// Mitsubishi GX Works2 project: 40国轩高温2次注液尝试优化   PLC: Q06UDEH

TYPE ConveyorIO : STRUCT
  xUnloadCCW : BOOL;  (* 下料为反转 *)
  xUnloadAlarm : BOOL;  (* 下料报警 *)
  xUnload : BOOL;  (* 下料请求 *)
  xPutInto : BOOL;  (* 线体直接投入物料 *)
  xNotArriveAlarm : BOOL;  (* 未到达报警 *)
  xNextRun : BOOL;  (* 下段线体运行 *)
  xMotorCW : BOOL;  (* 电机正转 *)
  xMotorCCW : BOOL;  (* 电机反转 *)
  xManual : BOOL;  (* 手动 *)
  xloadCCW : BOOL;  (* 上料为反转 *)
  xLimitAlarrm : BOOL;  (* 限位报警 *)
  xLoad : BOOL;  (* 上料请求 *)
  xForward : BOOL;  (* 正转手动 *)
  xEmpty : BOOL;  (* 线体状态为空 *)
  xCWPresent : BOOL;  (* 正转检测有无传感器 *)
  xCCWPresent : BOOL;  (* 反转检测有无传感器 *)
  xBusy : BOOL;  (* 工作中 *)
  xBackward : BOOL;  (* 反转手动 *)
  xAuto : BOOL;  (* 自动 *)
  xPosLimit : BOOL;  (* 正限位 *)
  xNegLimit : BOOL;  (* 负限位 *)
  xOverWidthAlarm : BOOL;  (* 超宽报警 *)
  xError : BOOL;  (* 报警 *)
  iProductCategoryIn : INT;  (* 产品类型输入 *)
  iProductCategory : INT;  (* 产品类型记录 *)
  iProductCategoryOut : INT;  (* 产品类型输出 *)
  diDeviceID : DINT;  (* 设备编号 *)
  tUnloadAlarmDelay : TIME;  (* 下料报警时间设置 *)
  tLoadDelay : TIME;  (* 上料延时设置 *)
  xSizeDeficientDetect : BOOL;  (* 尺寸缺陷检测 *)
  xZoneClear : BOOL;  (* 初始化线体清除 *)
  tZoneClearTime : TIME;  (* 初始化线体清除时间 *)
  iTaskIDIn : INT;  (* 产品类型输入 *)
  iTaskID : INT;  (* 产品类型记录 *)
  iTaskIDOut : INT;  (* 产品类型输出 *)
  diDesConveyorIn : DINT;  (* 产品类型输入 *)
  diDesConveyor : DINT;  (* 产品类型记录 *)
  diDesConveyorOut : DINT;  (* 产品类型输出 *)
END_STRUCT END_TYPE

TYPE ShuttleCarIO : STRUCT
  xReady : BOOL;  (* 准备就绪 *)
  xForward : BOOL;  (* 正转 *)
  xBackward : BOOL;  (* 反转 *)
  iCurrentPos : INT;  (* 当前位置 *)
  iDestinationPos : INT;  (* 目标位置 *)
  xCW : BOOL;  (* 正转输出 *)
  xCCW : BOOL;  (* 反转输出 *)
  xBrake : BOOL;  (* 刹车 *)
  xHomeSwitch : BOOL;  (* 零位接近开关 *)
  xPosLimit : BOOL;  (* 正限位 *)
  xNegLimit : BOOL;  (* 负限位 *)
  xMDIExe : BOOL;  (* MDI开始 *)
  xMDIDone : BOOL;  (* MDI 完成 *)
  xPassLimit : BOOL;  (* 限位屏蔽 *)
  xPosLimitCatch : BOOL;  (* 正限位捕捉 *)
  xNegLimitCatch : BOOL;  (* 负限位捕捉 *)
  xHomeExe : BOOL;  (* 开始寻零 *)
  xHomeDone : BOOL;  (* 寻零完成 *)
  xHomeBusy : BOOL;  (* 寻零中 *)
  xHomeFailed : BOOL;  (* 寻零失败 *)
  xBusy : BOOL;  (* 工作中 *)
  tArriveDelay : TIME;  (* 到位延时 *)
  xCylinder : BOOL;  (* 气缸控制 *)
  tBrakeDelay : TIME;  (* 抱闸延时 *)
  xPauseRamp : BOOL;  (* 暂停减速斜坡标志位 *)
  xPresentDetect1 : BOOL;  (* 物料有无检测1 *)
  xPresentDetect2 : BOOL;  (* 物料有无检测2 *)
  xOvertimeAlarm : BOOL;  (* 超时报警 *)
  tSetOverTime : TIME;  (* 设置超时时间 *)
  xLooseDetect : BOOL;  (* 松绳检测 *)
  xLooseAlarm : BOOL;  (* 松绳报警 *)
  xArrive : BOOL;  (* 到位信号 *)
  diDeviceID : DINT;  (* 设备编号 *)
  xMoveStep : BOOL;  (* 寸动 *)
  xAdrSwitch : ARRAY [1..8] OF BOOL;  (* 位置开关 *)
END_STRUCT END_TYPE

TYPE SwitchIO : STRUCT
  xLiftCylinderRetractDetect : BOOL;
  xLiftCylinderExtendDetect : BOOL;
  xLiftCylinderRetract : BOOL;
  xLiftCylinderExtend : BOOL;
  xEntryBarCylinderRetract : BOOL;
  xLiftCylinderExtendInit : BOOL;
  xEntryEnable : BOOL;
  xExitEnable : BOOL;
  xExitBarCylinderRetract : BOOL;
  xSwithEnable : BOOL;
  xLiftCylinderRetractButton : BOOL;
  xLiftCylinderExtendButton : BOOL;
  xEntryBarCylinderRetractButton : BOOL;
  xExitBarCylinderRetractButton : BOOL;
  xPutInto : BOOL;  (* 单体复位 *)
  tSetOvertime : TIME;  (* 设定超时报警时间 *)
  xOvertimeAlarm : BOOL;  (* 超时报警 *)
END_STRUCT END_TYPE

TYPE QueueElement : STRUCT
  xCondition : BOOL;
  iPriority : INT;
END_STRUCT END_TYPE

TYPE UConveyorIO : STRUCT
  xLiftCylinderRetractDetect1 : BOOL;
  xLiftCylinderRetractDetect2 : BOOL;
  xLiftCylinderExtendDetect1 : BOOL;
  xLiftCylinderExtendDetect2 : BOOL;
  xLiftCylinderRetract1 : BOOL;
  xLiftCylinderRetract2 : BOOL;
  xLiftCylinderExtend1 : BOOL;
  xLiftCylinderExtend2 : BOOL;
  xExitBarCylinderRetract1 : BOOL;
  xExitBarCylinderRetract2 : BOOL;
  xLiftCylinderExtendInit1 : BOOL;
  xLiftCylinderExtendInit2 : BOOL;
  xEntryEnable1 : BOOL;
  xEntryEnable2 : BOOL;
  xEntryEnable3 : BOOL;
  xExitEnable1 : BOOL;
  xExitEnable2 : BOOL;
  xExitEnable3 : BOOL;
  xPassEnable : BOOL;  (* 直接放行去下段 *)
  xLiftCylinderRetractButton1 : BOOL;
  xLiftCylinderRetractButton2 : BOOL;
  xLiftCylinderExtendButton1 : BOOL;
  xLiftCylinderExtendButton2 : BOOL;
  xExitBarCylinderRetractButton1 : BOOL;
  xExitBarCylinderRetractButton2 : BOOL;
  xPutInto : BOOL;  (* 单体复位 *)
  tSetOvertime : TIME;  (* 设定超时报警时间 *)
  xOvertimeAlarm : BOOL;  (* 超时报警 *)
  iTask : INT;  (* 3个任务 *)
  xBatteryDetect1 : BOOL;  (* 电池检测1 *)
  xBatteryDetect2 : BOOL;  (* 电池检测2 *)
  xBatteryError : BOOL;  (* 空框里有电池错误 *)
END_STRUCT END_TYPE

TYPE FolderIO : STRUCT
  o_xCylinderGrabExtend : BOOL;  (* 气缸夹紧 *)
  o_xCylinderGrabRetract : BOOL;  (* 气缸松开 *)
  i_xCylinderGrabExtendDetect : BOOL;  (* 夹紧检测 *)
  i_xCylinderGrabRetractDetect : BOOL;  (* 松开检测 *)
  o_xCylinderUpExtend : BOOL;  (* 上层伸出 *)
  o_xCylinderUpRetract : BOOL;  (* 上层缩回 *)
  i_xCylinderUpExtendDetect : BOOL;  (* 上层伸出检测 *)
  i_xCylinderUpRetractDetect : BOOL;  (* 上层缩回检测 *)
  o_xCylinderDownExtend : BOOL;  (* 下层伸出 *)
  o_xCylinderDownRetract : BOOL;  (* 下层缩回 *)
  i_xCylinderDownExtendDetect : BOOL;  (* 下层伸出检测 *)
  i_xCylinderDownRetractDetect : BOOL;  (* 下层缩回检测 *)
  i_xExitEnable : BOOL;  (* 下料信号 *)
  i_xEntryEnable : BOOL;  (* 上料信号 *)
  o_xEntryPermit : BOOL;  (* 允许上料(拆盘需要，叠盘不需要) *)
  i_iFloor : INT;  (* 层数 *)
  i_xCylinderGrabExtendButton : BOOL;  (* 气缸夹紧按钮 *)
  i_xCylinderGrabRetractButton : BOOL;  (* 气缸松开按钮 *)
  i_xCylinderUpExtendButton : BOOL;  (* 上层伸出按钮 *)
  i_xCylinderUpRetractButton : BOOL;  (* 上层缩回按钮 *)
  i_xCylinderDownExtendButton : BOOL;  (* 下层伸出按钮 *)
  i_xCylinderDownRetractButton : BOOL;  (* 下层缩回按钮 *)
  o_xDownCylinderError : BOOL;  (* 下层气缸层伸出未到达 *)
  o_xUpCylinderError : BOOL;  (* 上层气缸伸出未到达 *)
  o_xGrabCylinderError : BOOL;  (* 夹紧气缸伸出未到达 *)
  i_tSetOvertime : TIME;  (* 未到达计时 *)
END_STRUCT END_TYPE

TYPE CommunicationIO : STRUCT
  i_iResponsPCPLC : INT;  (* 上位机写入-请求确认 *)
  i_iTypeInfoPCPLC : INT;  (* 上位机写入-批次标识，是否同批次 *)
  i_iReadWriteFlagPCPLC : INT;  (* 上位机写入-读写标志位 *)
  i_iTaskProcessFlagPCPLC : INT;  (* 上位机写入-任务处理标志位 *)
  i_iCommandPCPLC : INT;  (* 上位机写入-命令字 *)
  i_iTaskIDPCPLC : INT;  (* 上位机写入-任务号 *)
  i_diDestinationDevicePCPLC : DINT;  (* 上位机写入-目标设备号 *)
  i_iProductIDPCPLC : INT;  (* 上位机写入-框码后4位 *)
  o_iRequestPLCPC : INT;  (* 上位机读取-请求状态 *)
  o_iForceInportPLCPC : INT;  (* 上位机读取-强制入库 *)
  o_iFolderNumberPLCPC : INT;  (* 上位机读取-叠盘数量 *)
  o_iEmptyPLCPC : INT;  (* 上位机读取-有料状态 *)
  o_iReadWriteFlagPLCPC : INT;  (* 上位机读取-读写标志位 *)
  o_iDeviceStatusPLCPC : INT;  (* 上位机读取-设备状态 *)
  o_iTaskIDPLCPC : INT;  (* 上位机读取-任务号 *)
  o_iProductIDPLCPC : INT;  (* 上位机读取-框码后4位 *)
  i_xExtraCondition : BOOL;  (* 发送请求时的额外条件,比如需要升降到位 *)
  i_xExportConveyor : BOOL;  (* 线体是出库线体还是入库线体 *)
  i_xImportConveyor : BOOL;  (* 入库线体 *)
END_STRUCT END_TYPE

// global labels: Global
VAR_GLOBAL
  g_xAuto AT M11 : BOOL;
  g_xAutoSwitch AT X1 : BOOL;  (* 手自动钥匙旋钮 *)
  g_xManual : BOOL;
  g_xEStop AT X0 : BOOL;
  g_xAlarm : BOOL;
  g_xMute : BOOL;
  g_xStackLampRed AT Y200 : BOOL;
  g_xStackLampAmber AT Y201 : BOOL;
  g_xStackLampGreen AT Y202 : BOOL;
  g_xStop AT X3 : BOOL;
  g_xPause AT M3 : BOOL;  (* 暂停 *)
  g_xAutoStart AT X2 : BOOL;
  g_xAutoLamp AT Y204 : BOOL;
  g_xRemoteAutoStart AT M0 : BOOL;
  g_iConveyorStatus AT D4 : INT;
  g_xBuzzer AT Y203 : BOOL;
  g_xRemoteAuto AT M10 : BOOL;
  g_xReset AT X4 : BOOL;
  g_xResetSingle AT M4 : BOOL;  (* 单线体复位 *)
  g_xInsertTask AT M5 : BOOL;  (* 插入任务 *)
  g_diInsertDesConveyor AT D8 : DINT;
  g_iInsertTaskID AT D2 : INT;  (* 插入任务号 *)
  g_iInsertCategory AT D6 : INT;
  g_iState AT D40 : INT;
  g_iLocalAutoStep : BOOL;
  g_diDeviceIDSelect AT D0 : DINT;
  g_xTcpFailed : BOOL;  (* 通讯失败 *)
  g_xPickOver : ARRAY [1..4] OF BOOL;  (* 注液机给我们的信号，待定 *)
  g_x36HourExport1Forbidden AT M2 : BOOL;  (* 36H出库禁止 *)
  g_xForceImport AT M1 : BOOL;  (* 强制入库 *)
END_VAR

// task Task_01 (event TRUE, interval 0, priority 31): POU, START, TCP

PROGRAM POU
VAR
  Conveyor40102 : Conveyor;
  Conveyor40104 : Conveyor;
  Conveyor40105 : Conveyor;
  Conveyor40106 : Conveyor;
  Conveyor40103 : Conveyor;
  Conveyor40107 : Conveyor;
  Conveyor40108 : Conveyor;
  Conveyor40101 : Conveyor;
  Conveyor40109 : Conveyor;
  Conveyor40110 : Conveyor;
  Conveyor40111 : Conveyor;
  Conveyor40113 : Conveyor;
  Conveyor40114 : Conveyor;
  Conveyor40115 : Conveyor;
  Conveyor40116 : Conveyor;
  Conveyor40117 : Conveyor;
  Conveyor40118 : Conveyor;
  Conveyor40119 : Conveyor;
  Conveyor40120 : Conveyor;
  Conveyor40122 : Conveyor;
  Conveyor40124 : Conveyor;
  Conveyor40126 : Conveyor;
  Conveyor40129 : Conveyor;
  Conveyor40131 : Conveyor;
  Conveyor40133 : Conveyor;
  Conveyor40136 : Conveyor;
  Conveyor40137 : Conveyor;
  Conveyor40138 : Conveyor;
  Conveyor40140 : Conveyor;
  Conveyor401021 : Conveyor;
  Conveyor401101 : Conveyor;
  ConveyorIO40101 : ConveyorIO;
  ConveyorIO40103 : ConveyorIO;
  ConveyorIO40104 : ConveyorIO;
  ConveyorIO40105 : ConveyorIO;
  ConveyorIO40106 : ConveyorIO;
  ConveyorIO40107 : ConveyorIO;
  ConveyorIO40108 : ConveyorIO;
  ConveyorIO40109 : ConveyorIO;
  ConveyorIO40110 : ConveyorIO;
  ConveyorIO40111 : ConveyorIO;
  ConveyorIO40112 : ConveyorIO;
  ConveyorIO40113 : ConveyorIO;
  ConveyorIO40114 : ConveyorIO;
  ConveyorIO40115 : ConveyorIO;
  ConveyorIO40116 : ConveyorIO;
  ConveyorIO40117 : ConveyorIO;
  ConveyorIO40118 : ConveyorIO;
  ConveyorIO40119 : ConveyorIO;
  ConveyorIO40122 : ConveyorIO;
  ConveyorIO40124 : ConveyorIO;
  ConveyorIO40126 : ConveyorIO;
  ConveyorIO40128 : ConveyorIO;
  ConveyorIO40131 : ConveyorIO;
  ConveyorIO40132 : ConveyorIO;
  ConveyorIO40133 : ConveyorIO;
  ConveyorIO40135 : ConveyorIO;
  ConveyorIO40136 : ConveyorIO;
  ConveyorIO40137 : ConveyorIO;
  ConveyorIO40140 : ConveyorIO;
  ConveyorIO401021 : ConveyorIO;
  ConveyorIO401101 : ConveyorIO;
  Lifter40202 : ShuttleCar;
  Lifter40203 : ShuttleCar;
  Lifter40204 : ShuttleCar;
  Lifter40206 : ShuttleCar;
  LifterIO40202 : ShuttleCarIO;
  LifterIO40203 : ShuttleCarIO;
  LifterIO40204 : ShuttleCarIO;
  LifterIO40206 : ShuttleCarIO;
  Switch40302 : Switch;
  Switch40303 : Switch;
  Switch40304 : Switch;
  Switch40306 : Switch;
  Switch40307 : Switch;
  Switch40308 : Switch;
  Switch40309 : Switch;
  SwitchIO40301 : SwitchIO;
  SwitchIO40302 : SwitchIO;
  SwitchIO40303 : SwitchIO;
  SwitchIO40304 : SwitchIO;
  SwitchIO40305 : SwitchIO;
  SwitchIO40306 : SwitchIO;
  SwitchIO40307 : SwitchIO;
  SwitchIO40308 : SwitchIO;
  SwitchIO40309 : SwitchIO;
  Folder40501 : Folder;
  FolderIO40501 : FolderIO;
  DivideFolder40502 : DivideFolder;
  DivideFolderIO40502 : FolderIO;
  ConveyorIO40129 : ConveyorIO;
  Conveyor40112 : Conveyor;
  ConveyorIO40138 : ConveyorIO;
  Conveyor40128 : Conveyor;
  Conveyor40135 : Conveyor;
  Conveyor401061 : Conveyor;
  Lifter40201 : ShuttleCar;
  LifterIO40201 : ShuttleCarIO;
  Switch40301 : Switch;
  Conveyor40132 : Conveyor;
  ConveyorIO40102 : ConveyorIO;
  ConveyorIO401061 : ConveyorIO;
  Lifter40205 : ShuttleCar;
  LifterIO40205 : ShuttleCarIO;
  Switch40305 : Switch;
  Switch40310 : Switch;
  Switch40311 : Switch;
  Switch40312 : Switch;
  SwitchIO40310 : SwitchIO;
  SwitchIO40311 : SwitchIO;
  SwitchIO40312 : SwitchIO;
  ComConveyor40140 : ConveyorCommunication;
  ComConveyor40209 : ConveyorCommunication;
  ComConveyor40111 : ConveyorCommunication;
  ComConveyor40104 : ConveyorCommunication;
  ComConveyor40105 : ConveyorCommunication;
  ComConveyorIO40140 : CommunicationIO;
  ComConveyorIO40209 : CommunicationIO;
  ComConveyorIO40111 : CommunicationIO;
  ComConveyorIO40104 : CommunicationIO;
  ComConveyorIO40105 : CommunicationIO;
  Task40105 : PriorityQueue;  (* 4个位置要料请求排队 *)
  TaskCondition40105 : ARRAY [1..13] OF QueueElement;  (* 4个位置要料请求排队 *)
  m_iTask40105 : INT;  (* 4个位置要料请求排队 *)
  m_xLoadPermit : ARRAY [1..4] OF BOOL;  (* 4个·位置的上料许可，用触摸屏控制 *)
  m_xPickStrat : ARRAY [1..4] OF BOOL;  (* 4个位置的开始取料信号，给到注液机器 *)
  m_xPickDone : ARRAY [1..4] OF BOOL;  (* 4个取料完毕信号，注液机给我们 *)
  Conveyor401131 : Conveyor;
  Conveyor401161 : Conveyor;
  Conveyor401191 : Conveyor;
  ConveyorIO40120 : ConveyorIO;
  ConveyorIO401161 : ConveyorIO;
  ConveyorIO401131 : ConveyorIO;
  ConveyorIO401191 : ConveyorIO;
  Lifter40207 : ShuttleCar;
  Lifter40208 : ShuttleCar;
  LifterIO40207 : ShuttleCarIO;
  LifterIO40208 : ShuttleCarIO;
  Conveyor40134 : Conveyor;
  ConveyorIO40134 : ConveyorIO;
  ConveyorIO40209 : ConveyorIO;
  Conveyor40209 : Conveyor;
  m_xImport : BOOL;  (* 高温房上料多转一会儿 *)
  m_xExport : BOOL;  (* 高温房下料多转一会儿 *)
  m_TonImportDelay : TON;  (* 高温房入库延时 *)
  m_xImportDelay : BOOL;  (* 高温房入库延时 *)
  m_tImportDelay : TIME;  (* 高温房入库延时 *)
  m_TonExportDelay : TON;  (* 高温房出库延时 *)
  m_xExportDelay : BOOL;  (* 高温房出库延时 *)
  m_tExportDelay : TIME;  (* 高温房出库延时 *)
  TaskSwitch40305 : PreemptivePriority;  (* 1线入口任务队列 *)
  TaskCondition40305 : ARRAY [1..13] OF BOOL;  (* 1线入口任务队列 *)
  m_iTask40305 : INT;  (* 1线入口任务队列 *)
  TaskSwitch40306 : PreemptivePriority;  (* 2线入口任务队列 *)
  TaskCondition40306 : ARRAY [1..13] OF BOOL;  (* 2线入口任务队列 *)
  m_iTask40306 : INT;  (* 2线入口任务队列 *)
  TaskSwitch40307 : PreemptivePriority;  (* 3线入口任务队列 *)
  TaskCondition40307 : ARRAY [1..13] OF BOOL;  (* 3线入口任务队列 *)
  m_iTask40307 : INT;  (* 3线入口任务队列 *)
END_VAR
(*与注液机对接信号*)(*
	Y205:=M700;
	Y206:=M701;
	Y207:=M702;
	Y239:=M703;
	M705:=X4A AND X4B AND X4C AND X4D;
	*)
	OUT_T(m_xPickStrat[1] AND g_xAuto , TC1 ,10 );
	OUT_T(m_xPickStrat[2] AND g_xAuto , TC2 ,10 );
	OUT_T(m_xPickStrat[3] AND g_xAuto , TC3 ,10 );
	OUT_T(m_xPickStrat[4] AND g_xAuto , TC4 ,10 );
	Y205:=TS1;(*他们要求到位延时1秒给信号*)
	Y206:=TS2;
	Y207:=TS3;
	Y239:=TS4;
	g_xPickOver[1]:=X4A;
	g_xPickOver[2]:=X4B;
	g_xPickOver[3]:=X4C;
	g_xPickOver[4]:=X4D;		
Conveyor40140(ConveyorMotor:=ConveyorIO40140);(*叠盘前，虚拟扫码工位*)														
ConveyorIO40140.diDeviceID:=40140;	
ConveyorIO40140.xCWPresent:=D421.7;(*不良品工位的光电*)
ConveyorIO40140.xPutInto:=D421.9;(*状态刷新*)

Conveyor40209(ConveyorMotor:=ConveyorIO40209);(*起始叠盘和高温入横向线体*)
ConveyorIO40209.xCWPresent:=X39;						
Y234:=ConveyorIO40209.xMotorCW OR ConveyorIO40101.xMotorCW;						
ConveyorIO40209.xForward:=M542;						
M339:= NOT ConveyorIO40209.xEmpty;						
M639:=ConveyorIO40209.xError;						
ConveyorIO40209.diDeviceID:=40209;	
ConveyorIO40209.tLoadDelay:=t#4000ms;

Conveyor40101(ConveyorMotor:=ConveyorIO40101);(*高温入库横向*)
ConveyorIO40101.xCWPresent:=X8;						
(*Y208:=ConveyorIO40101.xMotorCW;						
ConveyorIO40101.xForward:=M500;*)						
M301:= NOT ConveyorIO40101.xEmpty;						
M601:=ConveyorIO40101.xError;						
ConveyorIO40101.diDeviceID:=40101;						
ConveyorIO40101.tLoadDelay:=t#4000ms;

Conveyor40102(ConveyorMotor:=ConveyorIO40102);(*高温入库竖向*)
ConveyorIO40102.xCCWPresent:=X8;
Y209:=ConveyorIO40102.xMotorCW OR ConveyorIO401021.xMotorCW;						
ConveyorIO40102.xForward:=M501;						
M302:= NOT ConveyorIO401021.xEmpty;						
M602:=ConveyorIO40102.xError OR ConveyorIO401021.xError;						
ConveyorIO40102.diDeviceID:=401021;						

Conveyor401021(ConveyorMotor:=ConveyorIO401021);(*虚拟的，入库门前停止位*)
ConveyorIO401021.xCWPresent:=X9;						
ConveyorIO401021.diDeviceID:=40102;		

Conveyor40103(ConveyorMotor:=ConveyorIO40103);(*高温入库门后，竖向*)
ConveyorIO40103.xCWPresent:=XA OR X5;					
Y20A:=ConveyorIO40103.xMotorCW;						
ConveyorIO40103.xForward:=M502;						
M303:= NOT ConveyorIO40103.xEmpty;						
M603:=ConveyorIO40103.xError;						
ConveyorIO40103.diDeviceID:=40103;						
ConveyorIO40103.tLoadDelay:=t#4000ms;

Conveyor40104(ConveyorMotor:=ConveyorIO40104);(*高温入库后横向*)
ConveyorIO40104.xCWPresent:=XA OR X5;						
Y20B:=ConveyorIO40104.xMotorCW OR m_xImport;						
ConveyorIO40104.xForward:=M503;						
M304:= NOT ConveyorIO40104.xEmpty;						
M604:=ConveyorIO40104.xError;						
ConveyorIO40104.diDeviceID:=40104;	

Conveyor40111(ConveyorMotor:=ConveyorIO40111);(*高温入库对接线体*)										
ConveyorIO40111.xCWPresent:=X7E;						
Y212:=ConveyorIO40111.xMotorCW;						
ConveyorIO40111.xForward:=M510;						
M311:= NOT ConveyorIO40111.xEmpty;						
M611:=ConveyorIO40111.xError;						
ConveyorIO40111.diDeviceID:=40111;	
ConveyorIO40111.tLoadDelay:=t#2S;	

Conveyor40105(ConveyorMotor:=ConveyorIO40105);(*高温出库对接线体*)
ConveyorIO40105.xCWPresent:=X7B;						
Y20C:=ConveyorIO40105.xMotorCW;						
ConveyorIO40105.xForward:=M504;						
M305:= NOT ConveyorIO40105.xEmpty;						
M605:=ConveyorIO40105.xError;						
ConveyorIO40105.diDeviceID:=40105;						

Conveyor40108(ConveyorMotor:=ConveyorIO40108);(*高温出库里面横向*)
ConveyorIO40108.xCWPresent:=XF OR X7;						
Y20F:=ConveyorIO40108.xMotorCW OR m_xExport;						
ConveyorIO40108.xForward:=M507;						
M308:= NOT ConveyorIO40108.xEmpty;						
M608:=ConveyorIO40108.xError;						
ConveyorIO40108.diDeviceID:=40108;	
ConveyorIO40108.tLoadDelay:=T#4000MS;

Conveyor40107(ConveyorMotor:=ConveyorIO40107);(*高温出库，里面竖向*)
ConveyorIO40107.xCWPresent:=XF OR X7;						
Y20E:=ConveyorIO40107.xMotorCW OR ConveyorIO401061.xMotorCW;						
ConveyorIO40107.xForward:=M506;						
M307:= NOT ConveyorIO401061.xEmpty;						
M607:=ConveyorIO40107.xError OR ConveyorIO401061.xError;						
ConveyorIO40107.diDeviceID:=401061;		

Conveyor401061(ConveyorMotor:=ConveyorIO401061);(*出库门前停止位，虚拟一段*)
ConveyorIO401061.xCWPresent:=XE;										
ConveyorIO401061.diDeviceID:=40107;	

Conveyor40106(ConveyorMotor:=ConveyorIO40106);(*高温出库，外面竖向*)
ConveyorIO40106.xCWPresent:=XD;						
Y20D:=ConveyorIO40106.xMotorCW;						
ConveyorIO40106.xForward:=M505;						
M306:= NOT ConveyorIO40106.xEmpty;						
M606:=ConveyorIO40106.xError;						
ConveyorIO40106.diDeviceID:=40106;															
ConveyorIO40106.tLoadDelay:=T#4000MS;

Conveyor40109(ConveyorMotor:=ConveyorIO40109);(*高温出库横向,&拆盘机&1线横向*)
ConveyorIO40109.xCWPresent:=XD;						
Y224:=ConveyorIO40109.xMotorCW OR ConveyorIO40117.xMotorCW OR ConveyorIO40114.xMotorCW;						
ConveyorIO40109.xForward:=M508;						
M309:= NOT ConveyorIO40109.xEmpty;						
M609:=ConveyorIO40109.xError;						
ConveyorIO40109.diDeviceID:=40109;		

Conveyor40117(ConveyorMotor:=ConveyorIO40117);(*拆盘位置*)					
ConveyorIO40117.xCWPresent:=XC;									
ConveyorIO40117.xForward:=M516;						
M317:= NOT ConveyorIO40117.xEmpty;						
M617:=ConveyorIO40117.xError;						
ConveyorIO40117.diDeviceID:=40117;
ConveyorIO40117.tLoadDelay:=t#4000ms;

Conveyor40114(ConveyorMotor:=ConveyorIO40114);(*1线横向*)					
ConveyorIO40114.xCWPresent:=X10;											
M314:= NOT ConveyorIO40114.xEmpty;						
M614:=ConveyorIO40114.xError;						
ConveyorIO40114.diDeviceID:=40114;						
ConveyorIO40114.tLoadDelay:=T#2000MS;

Conveyor40110(ConveyorMotor:=ConveyorIO40110);(*1线入*)
ConveyorIO40110.xCWPresent:=X10;						
Y211:=ConveyorIO40110.xMotorCW OR ConveyorIO401101.xMotorCW;						
ConveyorIO40110.xForward:=M509;								
M610:=ConveyorIO40110.xError OR ConveyorIO401101.xError;						
ConveyorIO40110.diDeviceID:=401101;					

Conveyor401101(ConveyorMotor:=ConveyorIO401101);(*1线末端*)
ConveyorIO401101.xPosLimit:= X88;
ConveyorIO401101.xNegLimit:=X89;
ConveyorIO401101.xCWPresent:=X12;											
M310:= NOT ConveyorIO401101.xEmpty;			
ConveyorIO401101.diDeviceID:=40110;	
ConveyorIO401101.tLoadDelay:=t#1000ms;
Y278:=(g_xAuto AND NOT ConveyorIO401101.xEmpty AND NOT m_xPickDone[1] AND NOT M585)(*夹紧气缸*)
			OR(g_xManual AND M585);		(*AND NOT M585 临时这么改一下，因为他们测试阶段，需要人工拿走托盘，就要松开夹紧气缸*)
Y27F:=ConveyorIO401101.xNextRun OR (g_xManual AND M586);(*末端阻挡*)		

Conveyor40112(ConveyorMotor:=ConveyorIO40112);(*2线横向*)
ConveyorIO40112.xCWPresent:=X13;						
Y213:=ConveyorIO40112.xMotorCW;						
ConveyorIO40112.xForward:=M511;						
M312:= NOT ConveyorIO40112.xEmpty;						
M612:=ConveyorIO40112.xError;						
ConveyorIO40112.diDeviceID:=40112;						
ConveyorIO40112.tLoadDelay:=T#7500MS;


Conveyor40113(ConveyorMotor:=ConveyorIO40113);(*2线入*)
ConveyorIO40113.xCWPresent:=X13;						
Y214:=ConveyorIO40113.xMotorCW OR ConveyorIO401131.xMotorCW;						
ConveyorIO40113.xForward:=M512;											
M613:=ConveyorIO40113.xError OR ConveyorIO401131.xError;						
ConveyorIO40113.diDeviceID:=401131;										

Conveyor401131(ConveyorMotor:=ConveyorIO401131);(*2线末端*)
ConveyorIO401131.xPosLimit:= X8A;
ConveyorIO401131.xNegLimit:=X8B;
ConveyorIO401131.xCWPresent:=X15;											
M313:= NOT ConveyorIO401131.xEmpty;											
ConveyorIO401131.diDeviceID:=40113;	
ConveyorIO401131.tLoadDelay:=t#1000ms;
Y272:=(g_xAuto AND NOT ConveyorIO401131.xEmpty AND NOT m_xPickDone[2] AND NOT M587)(*夹紧气缸*)
			OR(g_xManual AND M587);		(*AND NOT M587 临时这么改一下，因为他们测试阶段，需要人工拿走托盘，就要松开夹紧气缸*)	
Y27E:=ConveyorIO401131.xNextRun OR (g_xManual AND M588);(*末端阻挡*)			

Conveyor40115(ConveyorMotor:=ConveyorIO40115);(*3线横向*)
ConveyorIO40115.xCWPresent:=X16;						
Y216:=ConveyorIO40115.xMotorCW;						
ConveyorIO40115.xForward:=M514;						
M315:= NOT ConveyorIO40115.xEmpty;						
M615:=ConveyorIO40115.xError;						
ConveyorIO40115.diDeviceID:=40115;						
ConveyorIO40115.tLoadDelay:=T#5000MS;

Conveyor40116(ConveyorMotor:=ConveyorIO40116)(*3线入*);
ConveyorIO40116.xCWPresent:=X16;						
Y217:=ConveyorIO40116.xMotorCW OR ConveyorIO401161.xMotorCW;						
ConveyorIO40116.xForward:=M515;											
M616:=ConveyorIO40116.xError OR ConveyorIO401161.xError;						
ConveyorIO40116.diDeviceID:=401161;								

Conveyor401161(ConveyorMotor:=ConveyorIO401161)(*3线末端*);
ConveyorIO401161.xPosLimit:=X8C;
ConveyorIO401191.xNegLimit:=X8D;
ConveyorIO401161.xCWPresent:=X18;									
M316:= NOT ConveyorIO401161.xEmpty;										
ConveyorIO401161.diDeviceID:=40116;	
ConveyorIO401161.tLoadDelay:=t#1000ms;
Y27D:=(g_xAuto AND NOT ConveyorIO401161.xEmpty AND NOT m_xPickDone[3] AND NOT M589)(*夹紧气缸*)
			OR(g_xManual AND M589);		(*AND NOT M587 临时这么改一下，因为他们测试阶段，需要人工拿走托盘，就要松开夹紧气缸*)	
Y274:=ConveyorIO401161.xNextRun OR (g_xManual AND M590);(*末端阻挡*)	

Conveyor40118(ConveyorMotor:=ConveyorIO40118);(*4线横向**)
ConveyorIO40118.xCWPresent:=X19;						
Y219:=ConveyorIO40118.xMotorCW;						
ConveyorIO40118.xForward:=M517;						
M318:= NOT ConveyorIO40118.xEmpty;						
M618:=ConveyorIO40118.xError;						
ConveyorIO40118.diDeviceID:=40118;						
ConveyorIO40118.tLoadDelay:=T#4000MS;

Conveyor40119(ConveyorMotor:=ConveyorIO40119);(*4线入*)
ConveyorIO40119.xCWPresent:=X19;						
Y21A:=ConveyorIO40119.xMotorCW OR ConveyorIO401191.xMotorCW;						
ConveyorIO40119.xForward:=M518;											
M619:=ConveyorIO40119.xError OR ConveyorIO40119.xError;						
ConveyorIO40119.diDeviceID:=401191;						

Conveyor401191(ConveyorMotor:=ConveyorIO401191);(*4线末端*)
ConveyorIO401191.xPosLimit:=1(*X1B*);
ConveyorIO401191.xNegLimit:=X93;
ConveyorIO401191.xCWPresent:=X92;											
M319:= NOT ConveyorIO401191.xEmpty;											
ConveyorIO401191.diDeviceID:=40119;
ConveyorIO401191.tLoadDelay:=t#1000ms;	
Y27C:=(g_xAuto AND NOT ConveyorIO401191.xEmpty AND NOT m_xPickDone[4] AND NOT M591)(*夹紧气缸*)
			OR(g_xManual AND M591);		(*AND NOT M587 临时这么改一下，因为他们测试阶段，需要人工拿走托盘，就要松开夹紧气缸*)	
Y245:=ConveyorIO401191.xNextRun OR (g_xManual AND M592);(*末端阻挡*)	


Conveyor40120(ConveyorMotor:=ConveyorIO40120);(*下层4横*)
(*ConveyorIO40120.xPosLimit:=X92;						
ConveyorIO40120.xNegLimit:=X93;		*)				
ConveyorIO40120.xCWPresent:=X1D;						
Y21E:=ConveyorIO40120.xMotorCW;						
ConveyorIO40120.xForward:=M519;						
M320:= NOT ConveyorIO40120.xEmpty;						
M620:=ConveyorIO40120.xError;						
ConveyorIO40120.diDeviceID:=40120;						
(*
Conveyor40121(ConveyorMotor:=ConveyorIO40121);
ConveyorIO40121.xCWPresent:=X1C;						
Y21C:=ConveyorIO40121.xMotorCW;						
ConveyorIO40121.xForward:=M520;						
M321:= NOT ConveyorIO40121.xEmpty;						
M621:=ConveyorIO40121.xError;						
ConveyorIO40121.diDeviceID:=40121;						
*)
Conveyor40122(ConveyorMotor:=ConveyorIO40122);(*下层4出*)
ConveyorIO40122.xCWPresent:=X1D;						
Y21D:=ConveyorIO40122.xMotorCW;						
ConveyorIO40122.xForward:=M521;						
M322:= NOT ConveyorIO40122.xEmpty;						
M622:=ConveyorIO40122.xError;						
ConveyorIO40122.diDeviceID:=40122;		
ConveyorIO40122.tLoadDelay:=T#4000MS;				
(*
Conveyor40123(ConveyorMotor:=ConveyorIO40123);
ConveyorIO40123.xCWPresent:=X1D;						
Y21E:=ConveyorIO40123.xMotorCW;						
ConveyorIO40123.xForward:=M522;						
M323:= NOT ConveyorIO40123.xEmpty;						
M623:=ConveyorIO40123.xError;						
ConveyorIO40123.diDeviceID:=40123;		*)				

Conveyor40124(ConveyorMotor:=ConveyorIO40124);(*下层3出*)
ConveyorIO40124.xCWPresent:=X20;						
Y21F:=ConveyorIO40124.xMotorCW;						
ConveyorIO40124.xForward:=M523;						
M324:= NOT ConveyorIO40124.xEmpty;						
M624:=ConveyorIO40124.xError;						
ConveyorIO40124.diDeviceID:=40124;		
ConveyorIO40124.tLoadDelay:=T#4000MS;				
(*
Conveyor40125(ConveyorMotor:=ConveyorIO40125);
ConveyorIO40125.xCWPresent:=X20;						
Y220:=ConveyorIO40125.xMotorCW;						
ConveyorIO40125.xForward:=M524;						
M325:= NOT ConveyorIO40125.xEmpty;						
M625:=ConveyorIO40125.xError;						
ConveyorIO40125.diDeviceID:=40125;						
*)
Conveyor40126(ConveyorMotor:=ConveyorIO40126);(*下层3横*)
ConveyorIO40126.xCWPresent:=X20;						
Y221:=ConveyorIO40126.xMotorCW;						
ConveyorIO40126.xForward:=M525;						
M326:= NOT ConveyorIO40126.xEmpty;						
M626:=ConveyorIO40126.xError;						
ConveyorIO40126.diDeviceID:=40126;									

Conveyor40128(ConveyorMotor:=ConveyorIO40128);(*下层2出*)
ConveyorIO40128.xCWPresent:=X23;						
Y223:=ConveyorIO40128.xMotorCW;						
ConveyorIO40128.xForward:=M527;						
M328:= NOT ConveyorIO40128.xEmpty;						
M628:=ConveyorIO40128.xError;						
ConveyorIO40128.diDeviceID:=40128;						
ConveyorIO40128.tLoadDelay:=T#4000MS;

Conveyor40129(ConveyorMotor:=ConveyorIO40129);(*下层2横*)
ConveyorIO40129.xCWPresent:=X23;						
Y210:=ConveyorIO40129.xMotorCW ;						
ConveyorIO40129.xForward:=M528;						
M329:= NOT ConveyorIO40129.xEmpty;						
M629:=ConveyorIO40129.xError;						
ConveyorIO40129.diDeviceID:=40129;						
(*
Conveyor40130(ConveyorMotor:=ConveyorIO40130);
ConveyorIO40130.xCWPresent:=X25;						
Y225:=ConveyorIO40130.xMotorCW;						
ConveyorIO40130.xForward:=M529;						
M330:= NOT ConveyorIO40130.xEmpty;						
M630:=ConveyorIO40130.xError;						
ConveyorIO40130.diDeviceID:=40130;*)						

Conveyor40131(ConveyorMotor:=ConveyorIO40131);(*下层1出*)
ConveyorIO40131.xCWPresent:=X26;						
Y226:=ConveyorIO40131.xMotorCW;						
ConveyorIO40131.xForward:=M530;						
M331:= NOT ConveyorIO40131.xEmpty;						
M631:=ConveyorIO40131.xError;						
ConveyorIO40131.diDeviceID:=40131;						
ConveyorIO40131.tLoadDelay:=T#4000MS;

Conveyor40132(ConveyorMotor:=ConveyorIO40132);(*下层1横*)
ConveyorIO40132.xCWPresent:=X26;						
Y227:=ConveyorIO40132.xMotorCW OR ConveyorIO40134.xMotorCW;						
ConveyorIO40132.xForward:=M531;											
M632:=ConveyorIO40132.xError OR ConveyorIO40134.xUnload;	
M332:= NOT ConveyorIO40132.xEmpty;						
ConveyorIO40132.diDeviceID:=40132;		
ConveyorIO40132.tLoadDelay:=t#4000ms;				

Conveyor40134(ConveyorMotor:=ConveyorIO40134);(*虚拟的，下层1横下一段*)
ConveyorIO40134.xCWPresent:=X27;																					
ConveyorIO40134.diDeviceID:=40134;		

Conveyor40133(ConveyorMotor:=ConveyorIO40133);(*下层输送*)
ConveyorIO40133.xCWPresent:=X28;						
Y228:=ConveyorIO40133.xMotorCW;						
ConveyorIO40133.xForward:=M532;						
M333:= NOT ConveyorIO40133.xEmpty;						
M633:=ConveyorIO40133.xError;						
ConveyorIO40133.diDeviceID:=40133;						
			

Conveyor40135(ConveyorMotor:=ConveyorIO40135);(*4线末端升降线体*)
(*ConveyorIO40135.xPosLimit:=X2C;						
ConveyorIO40135.xNegLimit:=X2B;	*)
ConveyorIO40135.xSizeDeficientDetect:=1;					
ConveyorIO40135.xCWPresent:=X2A;						
ConveyorIO40135.xCCWPresent:=X2B;						
Y22A:=ConveyorIO40135.xMotorCW;						
Y22B:=ConveyorIO40135.xMotorCCW;						
ConveyorIO40135.xForward:=M534;						
ConveyorIO40135.xBackward:=M535;						
M335:= NOT ConveyorIO40135.xEmpty;						
M635:=ConveyorIO40135.xError;						
ConveyorIO40135.diDeviceID:=40135;						

Conveyor40136(ConveyorMotor:=ConveyorIO40136);(*3线末端升降线体*)
(*ConveyorIO40136.xPosLimit:=X2F;						
ConveyorIO40136.xNegLimit:=X2E;		*)		
ConveyorIO40136.xSizeDeficientDetect:=1;		
ConveyorIO40136.xCWPresent:=X2d;						
ConveyorIO40136.xCCWPresent:=X2E;						
Y22D:=ConveyorIO40136.xMotorCW;						
Y22C:=ConveyorIO40136.xMotorCCW;						
ConveyorIO40136.xForward:=M536;						
ConveyorIO40136.xBackward:=M537;						
M336:= NOT ConveyorIO40136.xEmpty;						
M636:=ConveyorIO40136.xError;						
ConveyorIO40136.diDeviceID:=40136;						

Conveyor40137(ConveyorMotor:=ConveyorIO40137);(*2线末端升降线体*)
(*ConveyorIO40137.xPosLimit:=NOT X32;						
ConveyorIO40137.xNegLimit:=NOT X31;		*)		
ConveyorIO40137.xSizeDeficientDetect:=1;
ConveyorIO40137.xCWPresent:=X30;						
ConveyorIO40137.xCCWPresent:=X31;						
Y22E:=ConveyorIO40137.xMotorCW;						
Y22F:=ConveyorIO40137.xMotorCCW;						
ConveyorIO40137.xForward:=M538;						
ConveyorIO40137.xBackward:=M539;						
M337:= NOT ConveyorIO40137.xEmpty;						
M637:=ConveyorIO40137.xError;						
ConveyorIO40137.diDeviceID:=40137;						

Conveyor40138(ConveyorMotor:=ConveyorIO40138);(*1线末端升降线体*)
(*ConveyorIO40138.xPosLimit:=X35;						
ConveyorIO40138.xNegLimit:=X34;	*)	
ConveyorIO40138.xSizeDeficientDetect:=1;				
ConveyorIO40138.xCWPresent:=X33;						
ConveyorIO40138.xCCWPresent:=X83;						
Y231:=ConveyorIO40138.xMotorCW;						
Y230:=ConveyorIO40138.xMotorCCW;						
ConveyorIO40138.xForward:=M540;						
ConveyorIO40138.xBackward:=M541;						
M338:= NOT ConveyorIO40138.xEmpty;						
M638:=ConveyorIO40138.xError;						
ConveyorIO40138.diDeviceID:=40138;																					

Lifter40201(ShuttleCarInOut:=LifterIO40201);(*高温入库门*)
LifterIO40201.xCylinder:=1;
Y23A:=LifterIO40201.xCW;					
Y23B:=LifterIO40201.xCCW;					
LifterIO40201.xForward:=M543;					
LifterIO40201.xBackward:=M544;					
ShuttleCarCurrentPosition(X3F OR X3E,X3F,X3E,FALSE,LifterIO40201.iCurrentPos);					
M644:=LifterIO40201.xOvertimeAlarm ;					
LifterIO40201.diDeviceID:=40201;					

Lifter40202(ShuttleCarInOut:=LifterIO40202);		(*高温出库门*)
LifterIO40202.xCylinder:=1;			
Y23C:=LifterIO40202.xCW;					
Y23D:=LifterIO40202.xCCW;					
LifterIO40202.xForward:=M545;					
LifterIO40202.xBackward:=M546;					
ShuttleCarCurrentPosition(X41 OR X40,X41,X40,FALSE,LifterIO40202.iCurrentPos);					
M645:=LifterIO40202.xOvertimeAlarm ;					
LifterIO40202.diDeviceID:=40202;					

Lifter40203(ShuttleCarInOut:=LifterIO40203);		(*1线升降台*)
LifterIO40203.xCylinder:=1;			
Y23E:=LifterIO40203.xCW;					
Y23F:=LifterIO40203.xCCW;					
LifterIO40203.xForward:=M547;					
LifterIO40203.xBackward:=M548;					
ShuttleCarCurrentPosition(X43 OR X42,X42,X43,FALSE,LifterIO40203.iCurrentPos);					
M646:=LifterIO40203.xOvertimeAlarm ;					
LifterIO40203.diDeviceID:=40203;					